(* Logix 5000 project; controller MV vendor 1 type 14 code 217 rev 31.11; software revision 31.00; part 8 of 53 *)
(* tags used below, declared in another part *)
   CWD : CHECKWORD_FLAGS;
   MC_B240 : INT[255];   // CH1 RN PMP Channel 1 return pum p drive flags
   MC_B242 : INT[255];   // CH1 ROUTE Channel 1 route requ est flags
   MC_bit_returned : BOOL;
   MC_CH1_DR1 : PlantItem;   // CH1_DR1
   MC_CH1_DR2 : PlantItem;   // CH1_DR2
   MC_CH1_DT1 : PlantItem;   // CH1_DT1
   MC_CH1_DT2 : PlantItem;   // CH1_DT2
   MC_CH1_R1 : PlantItem;   // CH1_R1
   MC_CH1_R1R : PlantItem;   // CH1_R1R
   MC_CH1_R2 : PlantItem;   // CH1_R2
   MC_CH1_R2R : PlantItem;   // CH1_R2R
   MC_CH1_R3 : PlantItem;   // CH1_R3
   MC_CH1_R3R : PlantItem;   // CH1_R3R
   MC_CH1_R4 : PlantItem;   // CH1_R4
   MC_CH1_R4R : PlantItem;   // CH1_R4R
   MC_CH1_R5 : PlantItem;   // CH1_R5
   MC_CH1_R5R : PlantItem;   // CH1_R5R
   MC_CH1_R6 : PlantItem;   // CH1_R6
   MC_CH1_R6R : PlantItem;   // CH1_R6R
   MC_CH1_T105_2_ACC : DINT;
   MC_data_file_value_to_move : DINT;
   MC_N10 : INT[255];   // SETTINGS
   MC_N100 : INT[255];   // C1_PLC Channel 1 PLC data
   MC_N100_29_0_Storagebit : BOOL;
   MC_N102 : INT[255];   // CH1 PROG Channel 1 CIP progra m
   MC_N104 : INT[255];   // CH1 REPORT Channel 1 CIP report file
   MC_N112 : INT[255];   // FVR DATA Data read from FV ro uting PLC
   MC_N113 : INT[255];   // MVR DATA Data read from MV ro uting PLC
   MC_N114 : INT[255];   // YP DATA
   MC_N200 : INT[255];   // CHK_WORK Plant item fault che cking work area
   MC_N7 : INT[255];   // INTEGER
   MC_P1 : PlantItem;   // P1
   MC_PX_100 : PlantItem;   // PX_100
   MC_PX_101 : PlantItem;   // PX_101
   MC_T105 : TIMER[255];   // CH1 TIMERS Channel 1 timers
   MC_T4 : TIMER[255];   // TIMER
(* MC_Common, continued *)

ROUTINE MC_CH1_GLOBL_105   (* ladder *)
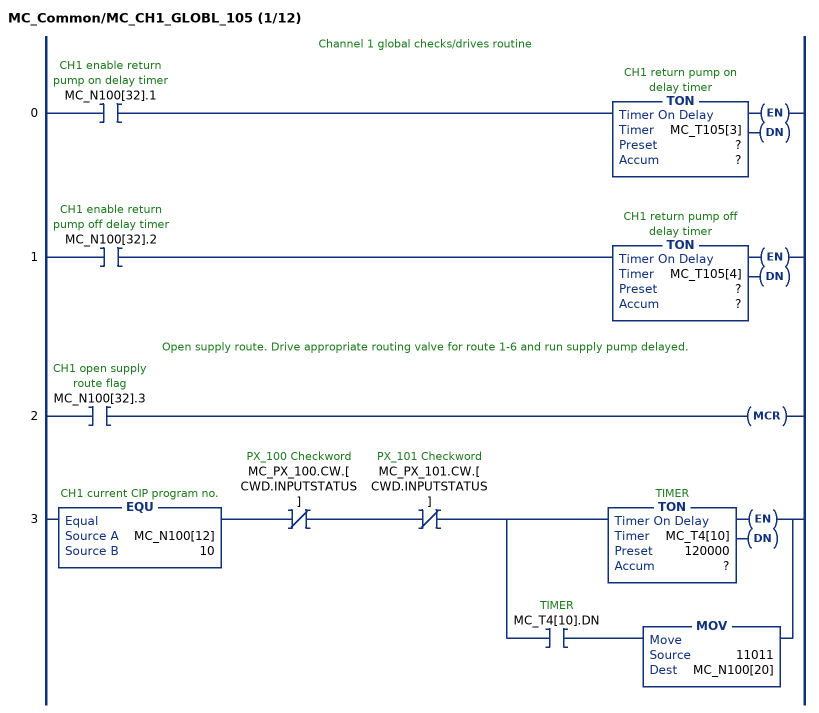
   // Channel 1 global checks/drives routine
   0: XIC(MC_N100[32].1)TON(MC_T105[3],?,?);
   1: XIC(MC_N100[32].2)TON(MC_T105[4],?,?);
   // Open supply route. Drive appropriate routing valve for route 1-6 and run supply pump delayed.
   2: XIC(MC_N100[32].3)MCR();
   3: EQU(MC_N100[12],10)XIO(MC_PX_100.CW.[CWD.INPUTSTATUS])XIO(MC_PX_101.CW.[CWD.INPUTSTATUS])[TON(MC_T4[10],?,?) ,XIC(MC_T4[10].DN) MOV(11011,MC_N100[20]) ];
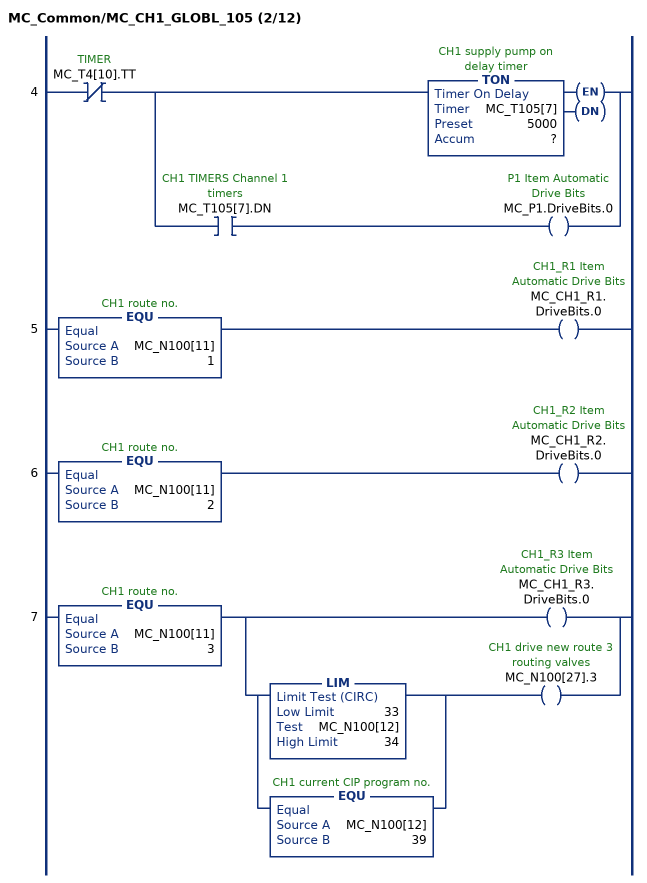
   4: XIO(MC_T4[10].TT)[TON(MC_T105[7],?,?) ,XIC(MC_T105[7].DN) OTE(MC_P1.DriveBits.0) ];
   5: EQU(MC_N100[11],1)OTE(MC_CH1_R1.DriveBits.0);
   6: EQU(MC_N100[11],2)OTE(MC_CH1_R2.DriveBits.0);
   7: EQU(MC_N100[11],3)[OTE(MC_CH1_R3.DriveBits.0) ,[LIM(33,MC_N100[12],34) ,EQU(MC_N100[12],39) ] OTE(MC_N100[27].3) ];
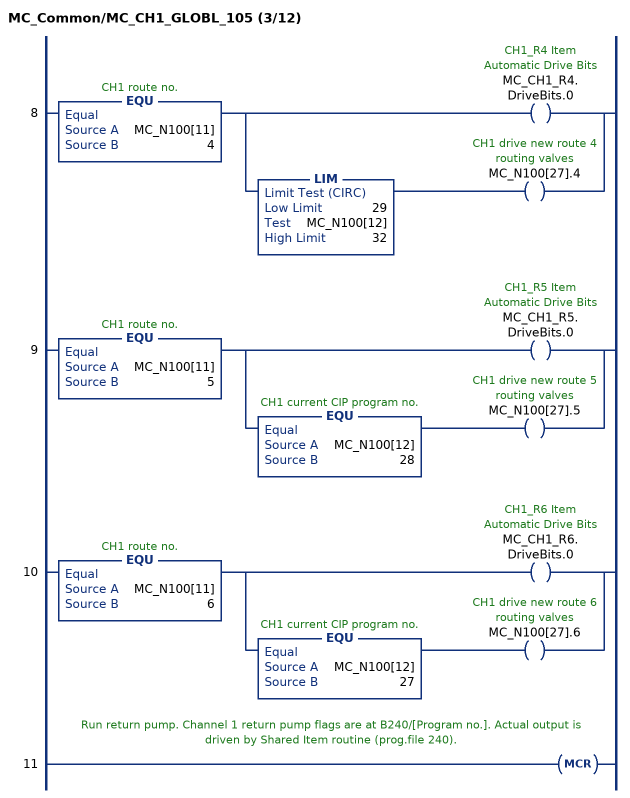
   8: EQU(MC_N100[11],4)[OTE(MC_CH1_R4.DriveBits.0) ,LIM(29,MC_N100[12],32) OTE(MC_N100[27].4) ];
   9: EQU(MC_N100[11],5)[OTE(MC_CH1_R5.DriveBits.0) ,EQU(MC_N100[12],28) OTE(MC_N100[27].5) ];
   10: EQU(MC_N100[11],6)[OTE(MC_CH1_R6.DriveBits.0) ,EQU(MC_N100[12],27) OTE(MC_N100[27].6) ];
   // Run return pump. Channel 1 return pump flags are at B240/[Program no.]. Actual output is driven by Shared Item routine (prog.file 240).
   11: MCR();
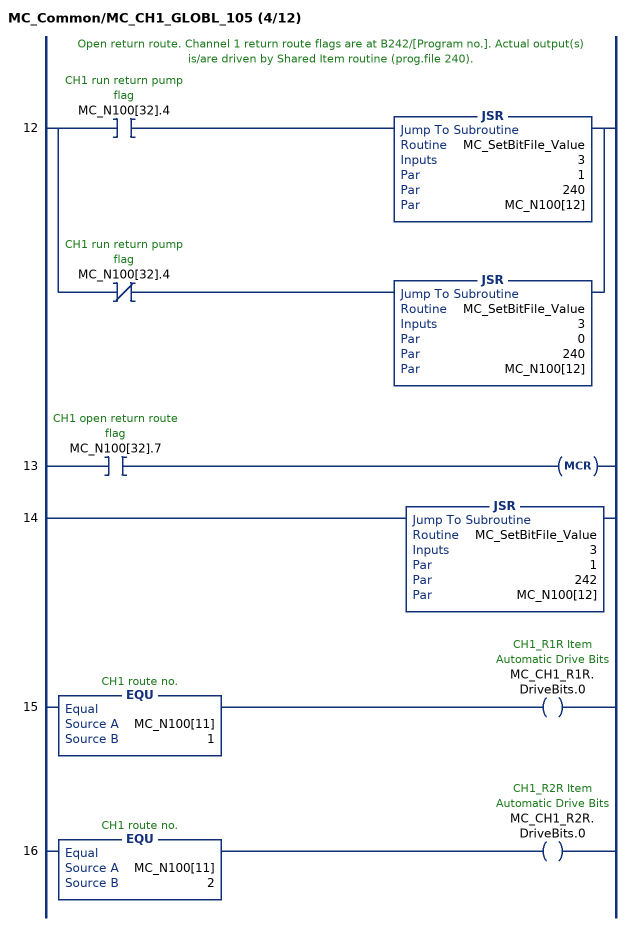
   // Open return route. Channel 1 return route flags are at B242/[Program no.]. Actual output(s) is/are driven by Shared Item routine (prog.file 240).
   12: [XIC(MC_N100[32].4) JSR(MC_SetBitFile_Value,3,1,240,MC_N100[12]) ,XIO(MC_N100[32].4) JSR(MC_SetBitFile_Value,3,0,240,MC_N100[12]) ];
   13: XIC(MC_N100[32].7)MCR();
   14: JSR(MC_SetBitFile_Value,3,1,242,MC_N100[12]);
   15: EQU(MC_N100[11],1)OTE(MC_CH1_R1R.DriveBits.0);
   16: EQU(MC_N100[11],2)OTE(MC_CH1_R2R.DriveBits.0);
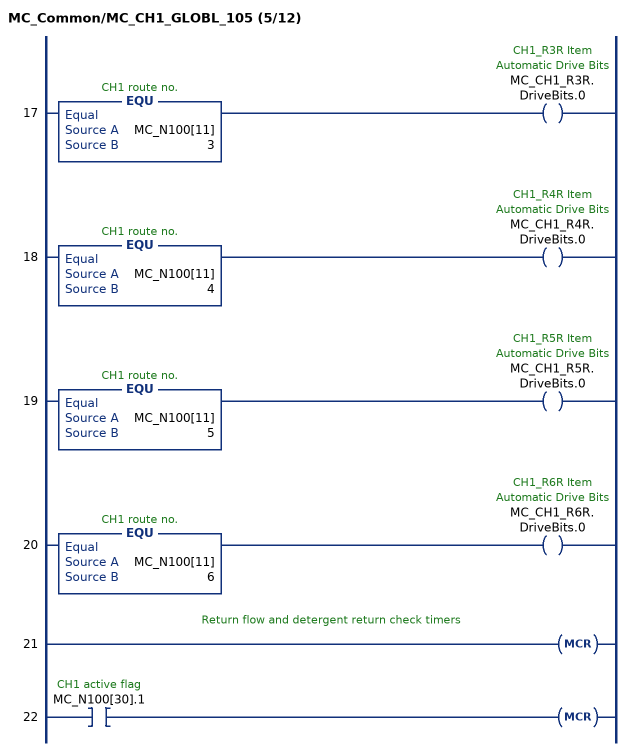
   17: EQU(MC_N100[11],3)OTE(MC_CH1_R3R.DriveBits.0);
   18: EQU(MC_N100[11],4)OTE(MC_CH1_R4R.DriveBits.0);
   19: EQU(MC_N100[11],5)OTE(MC_CH1_R5R.DriveBits.0);
   20: EQU(MC_N100[11],6)OTE(MC_CH1_R6R.DriveBits.0);
   // Return flow and detergent return check timers
   21: MCR();
   22: XIC(MC_N100[30].1)MCR();
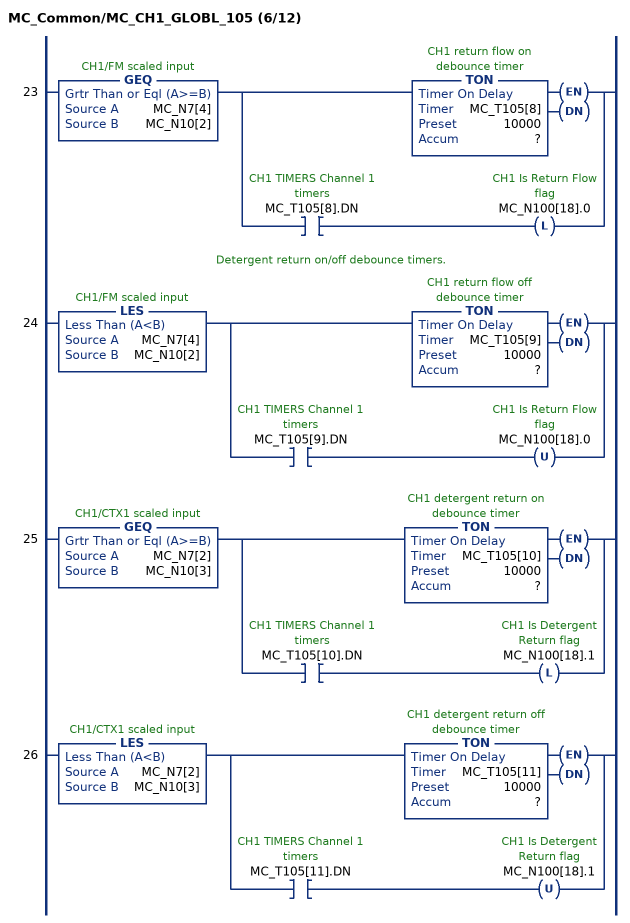
   23: GEQ(MC_N7[4],MC_N10[2])[TON(MC_T105[8],?,?) ,XIC(MC_T105[8].DN) OTL(MC_N100[18].0) ];
   // Detergent return on/off debounce timers.
   24: LES(MC_N7[4],MC_N10[2])[TON(MC_T105[9],?,?) ,XIC(MC_T105[9].DN) OTU(MC_N100[18].0) ];
   25: GEQ(MC_N7[2],MC_N10[3])[TON(MC_T105[10],?,?) ,XIC(MC_T105[10].DN) OTL(MC_N100[18].1) ];
   26: LES(MC_N7[2],MC_N10[3])[TON(MC_T105[11],?,?) ,XIC(MC_T105[11].DN) OTU(MC_N100[18].1) ];
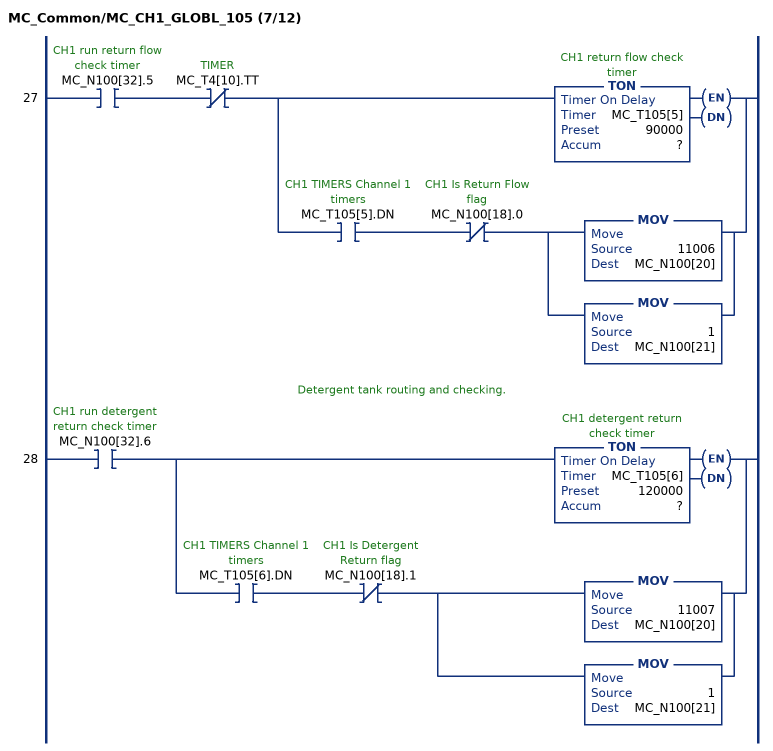
   27: XIC(MC_N100[32].5)XIO(MC_T4[10].TT)[TON(MC_T105[5],?,?) ,XIC(MC_T105[5].DN) XIO(MC_N100[18].0) [MOV(11006,MC_N100[20]) ,MOV(1,MC_N100[21]) ] ];
   // Detergent tank routing and checking.
   28: XIC(MC_N100[32].6)[TON(MC_T105[6],?,?) ,XIC(MC_T105[6].DN) XIO(MC_N100[18].1) [MOV(11007,MC_N100[20]) ,MOV(1,MC_N100[21]) ] ];
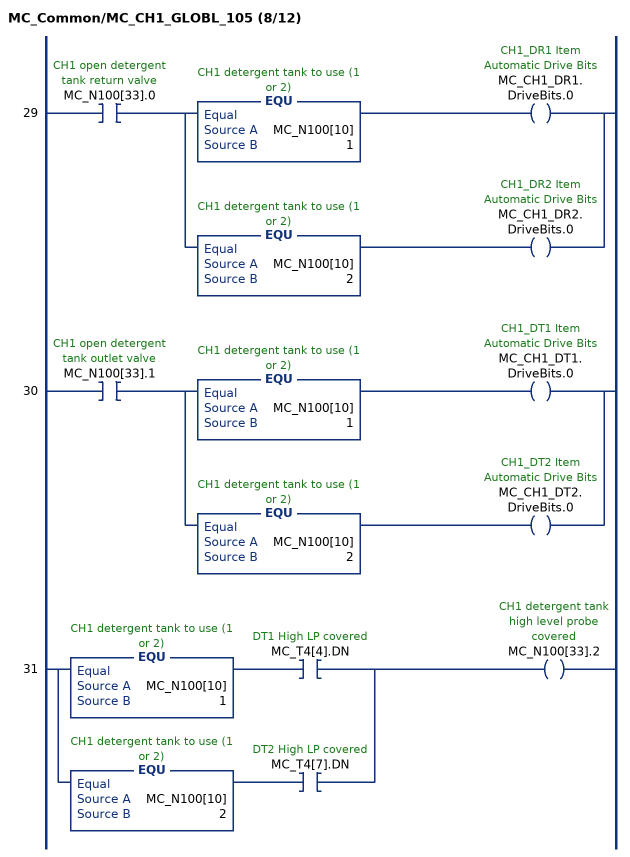
   29: XIC(MC_N100[33].0)[EQU(MC_N100[10],1) OTE(MC_CH1_DR1.DriveBits.0) ,EQU(MC_N100[10],2) OTE(MC_CH1_DR2.DriveBits.0) ];
   30: XIC(MC_N100[33].1)[EQU(MC_N100[10],1) OTE(MC_CH1_DT1.DriveBits.0) ,EQU(MC_N100[10],2) OTE(MC_CH1_DT2.DriveBits.0) ];
   31: [EQU(MC_N100[10],1) XIC(MC_T4[4].DN) ,EQU(MC_N100[10],2) XIC(MC_T4[7].DN) ]OTE(MC_N100[33].2);
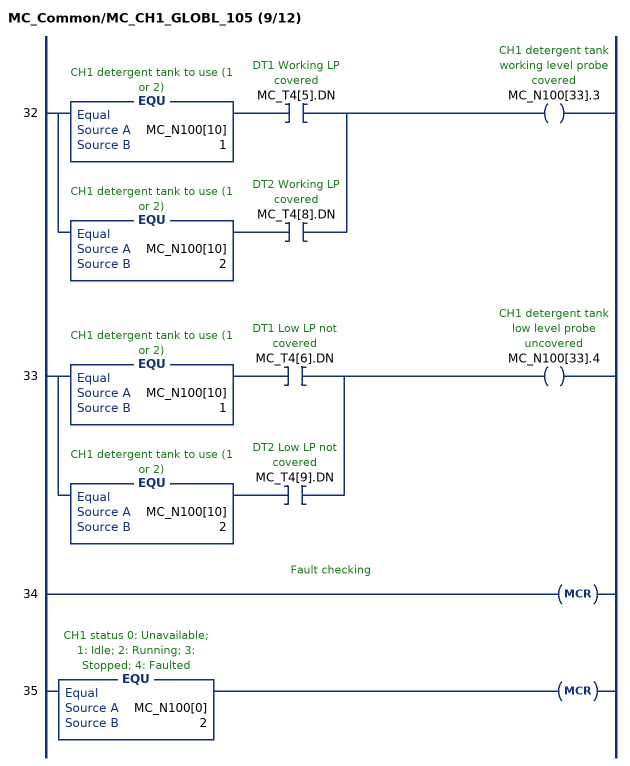
   32: [EQU(MC_N100[10],1) XIC(MC_T4[5].DN) ,EQU(MC_N100[10],2) XIC(MC_T4[8].DN) ]OTE(MC_N100[33].3);
   33: [EQU(MC_N100[10],1) XIC(MC_T4[6].DN) ,EQU(MC_N100[10],2) XIC(MC_T4[9].DN) ]OTE(MC_N100[33].4);
   // Fault checking
   34: MCR();
   35: EQU(MC_N100[0],2)MCR();
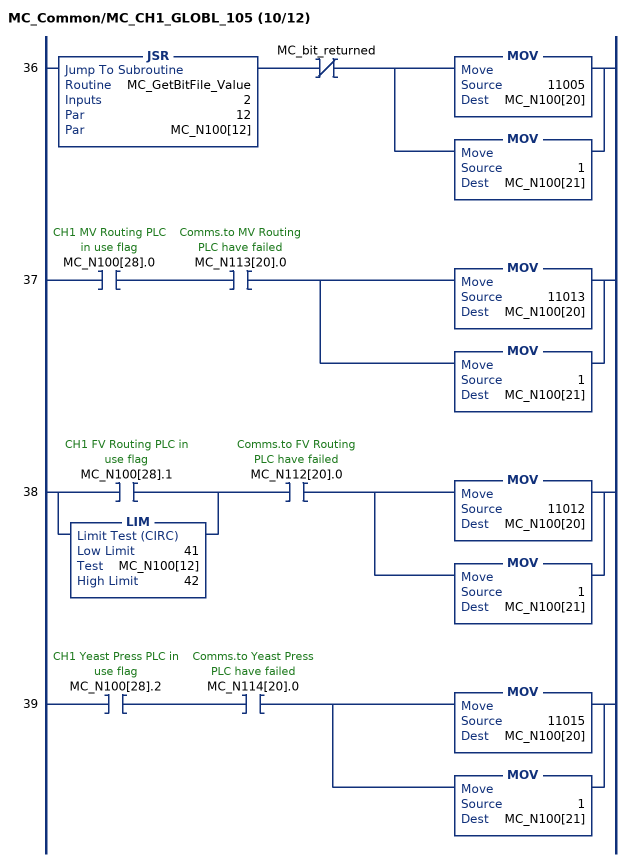
   36: JSR(MC_GetBitFile_Value,2,12,MC_N100[12])XIO(MC_bit_returned)[MOV(11005,MC_N100[20]) ,MOV(1,MC_N100[21]) ];
   37: XIC(MC_N100[28].0)XIC(MC_N113[20].0)[MOV(11013,MC_N100[20]) ,MOV(1,MC_N100[21]) ];
   38: [XIC(MC_N100[28].1) ,LIM(41,MC_N100[12],42) ]XIC(MC_N112[20].0)[MOV(11012,MC_N100[20]) ,MOV(1,MC_N100[21]) ];
   39: XIC(MC_N100[28].2)XIC(MC_N114[20].0)[MOV(11015,MC_N100[20]) ,MOV(1,MC_N100[21]) ];
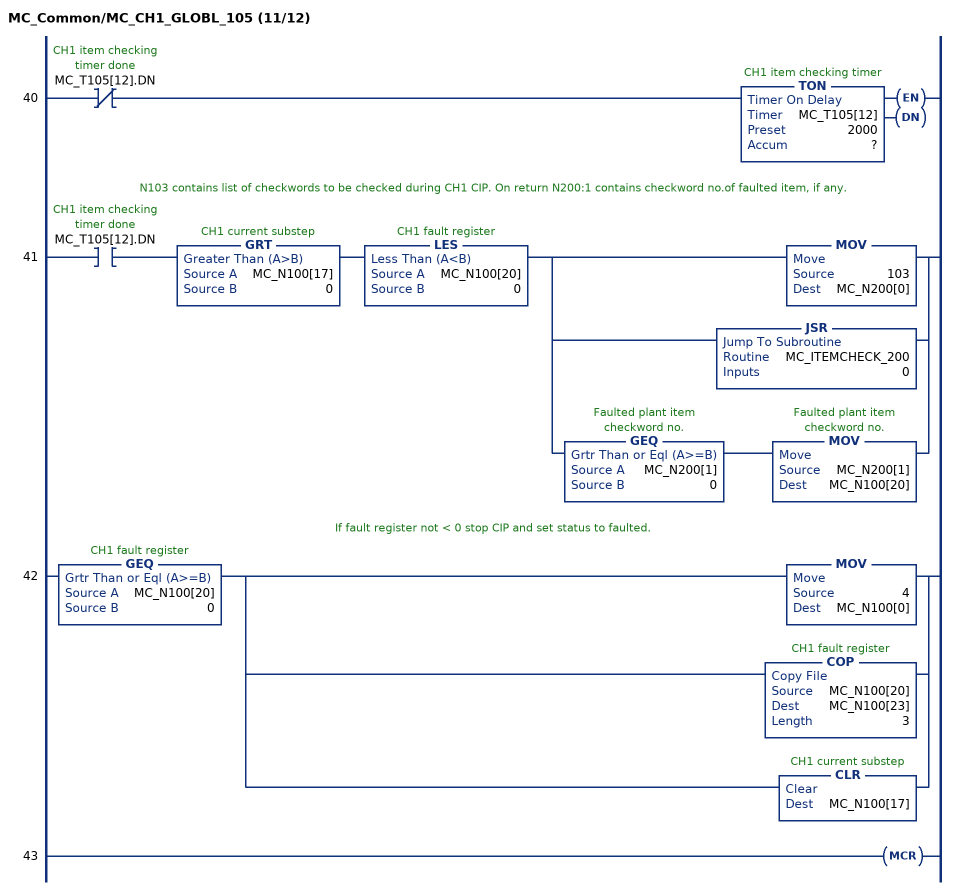
   40: XIO(MC_T105[12].DN)TON(MC_T105[12],?,?);
   // N103 contains list of checkwords to be checked during CH1 CIP. On return N200:1 contains checkword no.of faulted item, if any.
   41: XIC(MC_T105[12].DN)GRT(MC_N100[17],0)LES(MC_N100[20],0)[MOV(103,MC_N200[0]) ,JSR(MC_ITEMCHECK_200,0) ,GEQ(MC_N200[1],0) MOV(MC_N200[1],MC_N100[20]) ];
   // If fault register not < 0 stop CIP and set status to faulted.
   42: GEQ(MC_N100[20],0)[MOV(4,MC_N100[0]) ,COP(MC_N100[20],MC_N100[23],3) ,CLR(MC_N100[17]) ];
   43: MCR();
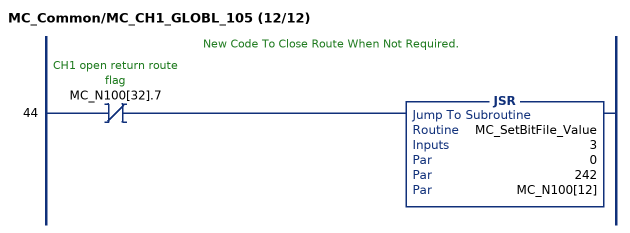
   // New Code To Close Route When Not Required.
   44: XIO(MC_N100[32].7)JSR(MC_SetBitFile_Value,3,0,242,MC_N100[12]);
END_ROUTINE

ROUTINE MC_CH1_MCP_100   (* ladder *)
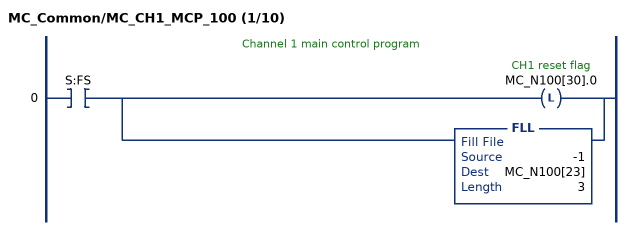
   // Channel 1 main control program
   0: XIC(S:FS)[OTL(MC_N100[30].0) ,FLL(-1,MC_N100[23],3) ];
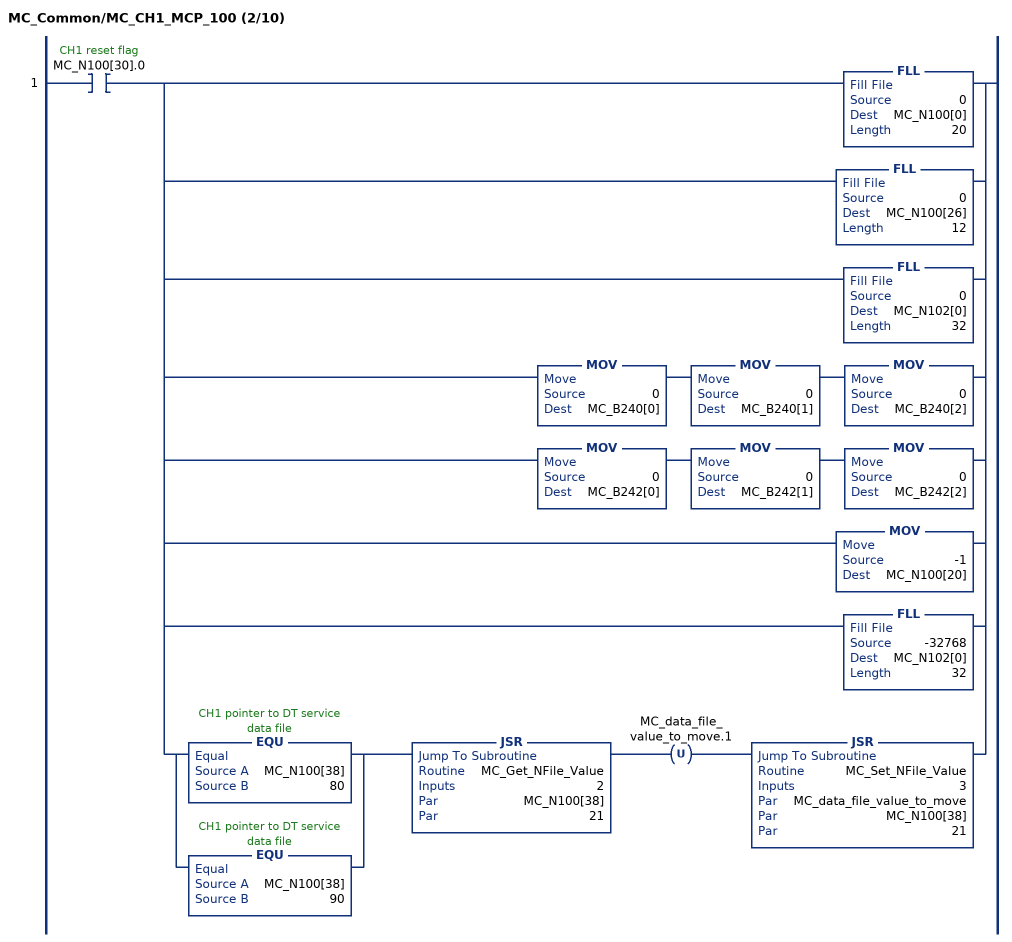
   1: XIC(MC_N100[30].0)[FLL(0,MC_N100[0],20) ,FLL(0,MC_N100[26],12) ,FLL(0,MC_N102[0],32) ,MOV(0,MC_B240[0]) MOV(0,MC_B240[1]) MOV(0,MC_B240[2]) ,MOV(0,MC_B242[0]) MOV(0,MC_B242[1]) MOV(0,MC_B242[2]) ,MOV(-1,MC_N100[20]) ,FLL(-32768,MC_N102[0],32) ,[EQU(MC_N100[38],80) ,EQU(MC_N100[38],90) ] JSR(MC_Get_NFile_Value,2,MC_N100[38],21) OTU(MC_data_file_value_to_move.1) JSR(MC_Set_NFile_Value,3,MC_data_file_value_to_move,MC_N100[38],21) ];
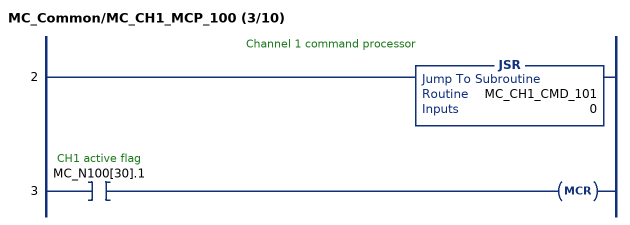
   // Channel 1 command processor
   2: JSR(MC_CH1_CMD_101,0);
   3: XIC(MC_N100[30].1)MCR();
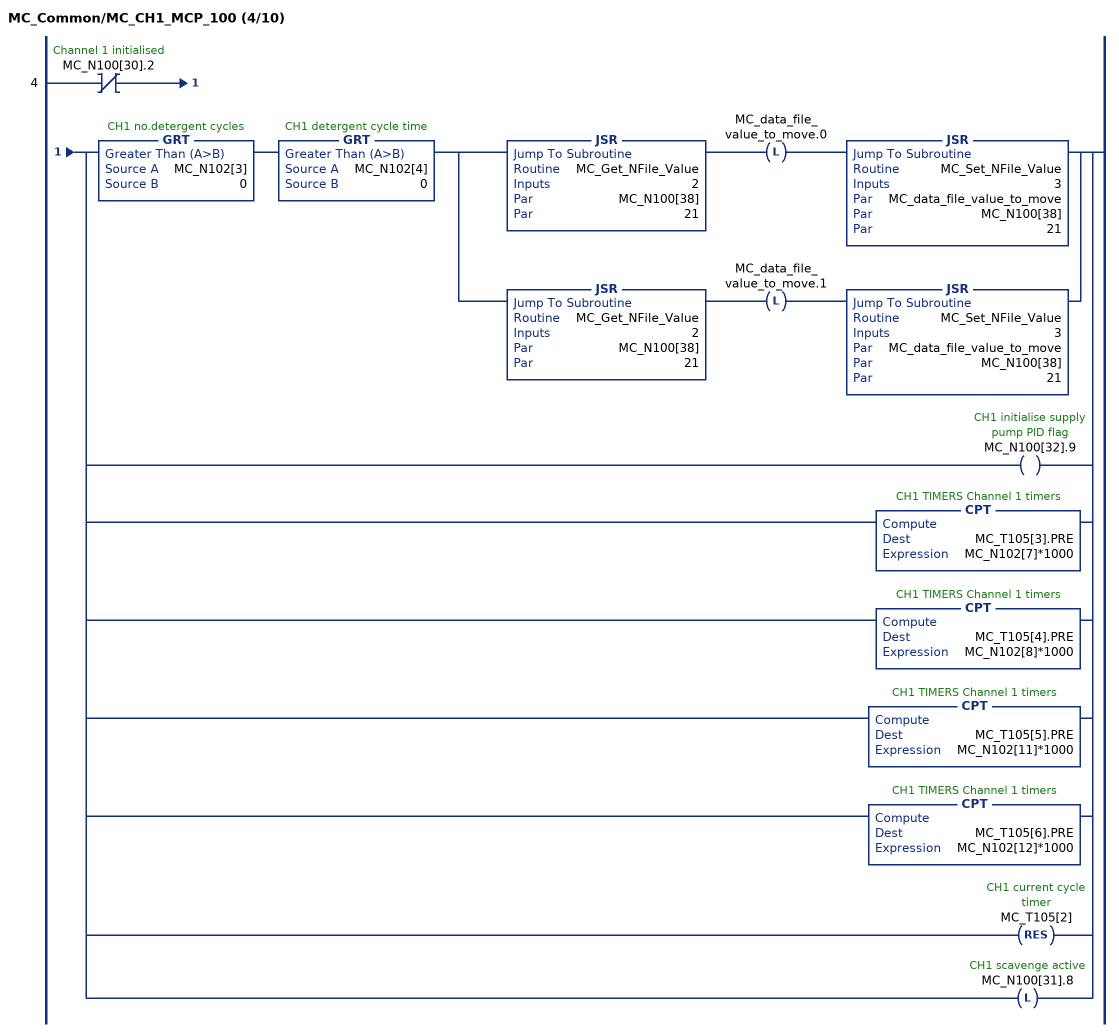
   4: XIO(MC_N100[30].2)[GRT(MC_N102[3],0) GRT(MC_N102[4],0) [JSR(MC_Get_NFile_Value,2,MC_N100[38],21) OTL(MC_data_file_value_to_move.0) JSR(MC_Set_NFile_Value,3,MC_data_file_value_to_move,MC_N100[38],21) ,JSR(MC_Get_NFile_Value,2,MC_N100[38],21) OTL(MC_data_file_value_to_move.1) JSR(MC_Set_NFile_Value,3,MC_data_file_value_to_move,MC_N100[38],21) ] ,OTE(MC_N100[32].9) ,[CPT(MC_T105[3].PRE,MC_N102[7]*1000) ,CPT(MC_T105[4].PRE,MC_N102[8]*1000) ,CPT(MC_T105[5].PRE,MC_N102[11]*1000) ,CPT(MC_T105[6].PRE,MC_N102[12]*1000) ,RES(MC_T105[2]) ,OTL(MC_N100[31].8) ] ];
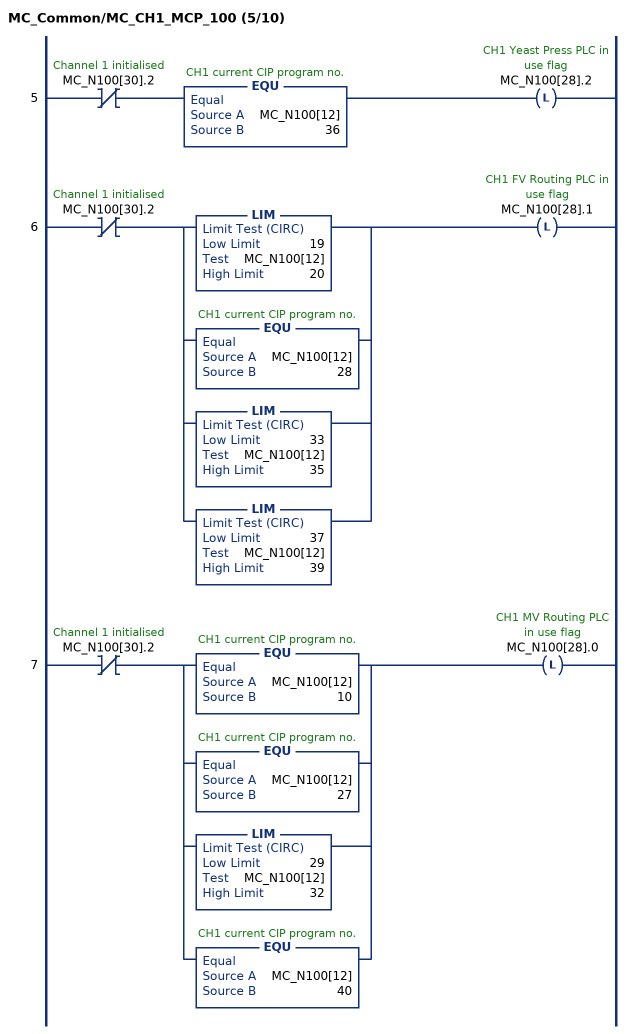
   5: XIO(MC_N100[30].2)EQU(MC_N100[12],36)OTL(MC_N100[28].2);
   6: XIO(MC_N100[30].2)[LIM(19,MC_N100[12],20) ,EQU(MC_N100[12],28) ,LIM(33,MC_N100[12],35) ,LIM(37,MC_N100[12],39) ]OTL(MC_N100[28].1);
   7: XIO(MC_N100[30].2)[EQU(MC_N100[12],10) ,EQU(MC_N100[12],27) ,LIM(29,MC_N100[12],32) ,EQU(MC_N100[12],40) ]OTL(MC_N100[28].0);
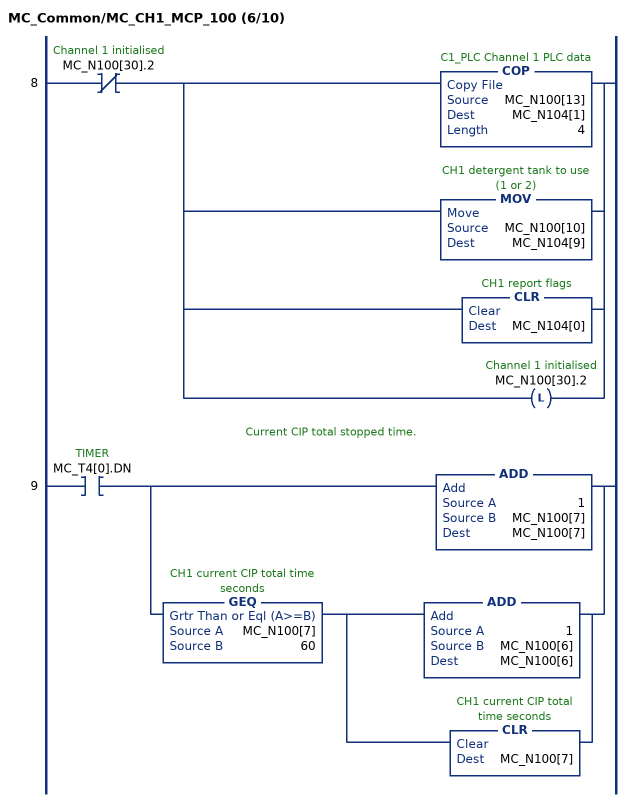
   8: XIO(MC_N100[30].2)[COP(MC_N100[13],MC_N104[1],4) ,MOV(MC_N100[10],MC_N104[9]) ,CLR(MC_N104[0]) ,OTL(MC_N100[30].2) ];
   // Current CIP total stopped time.
   9: XIC(MC_T4[0].DN)[ADD(1,MC_N100[7],MC_N100[7]) ,GEQ(MC_N100[7],60) [ADD(1,MC_N100[6],MC_N100[6]) ,CLR(MC_N100[7]) ] ];
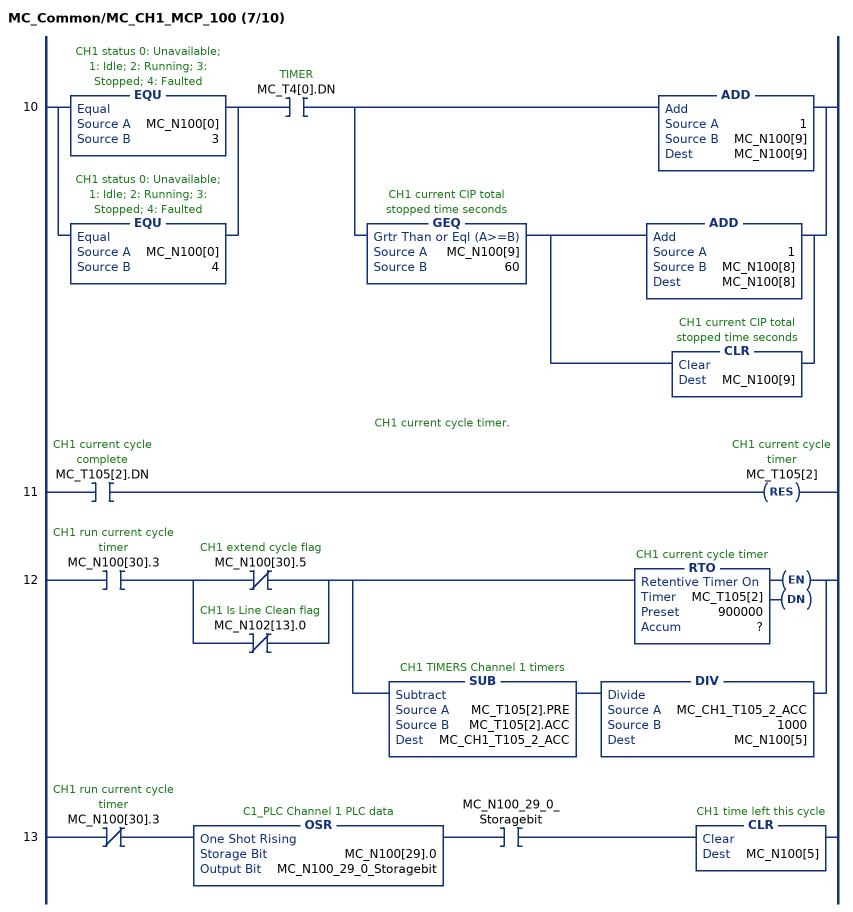
   10: [EQU(MC_N100[0],3) ,EQU(MC_N100[0],4) ]XIC(MC_T4[0].DN)[ADD(1,MC_N100[9],MC_N100[9]) ,GEQ(MC_N100[9],60) [ADD(1,MC_N100[8],MC_N100[8]) ,CLR(MC_N100[9]) ] ];
   // CH1 current cycle timer.
   11: XIC(MC_T105[2].DN)RES(MC_T105[2]);
   12: XIC(MC_N100[30].3)[XIO(MC_N100[30].5) ,XIO(MC_N102[13].0) ][RTO(MC_T105[2],?,?) ,SUB(MC_T105[2].PRE,MC_T105[2].ACC,MC_CH1_T105_2_ACC) DIV(MC_CH1_T105_2_ACC,1000,MC_N100[5]) ];
   13: XIO(MC_N100[30].3)OSR(MC_N100[29].0,MC_N100_29_0_Storagebit)XIC(MC_N100_29_0_Storagebit)CLR(MC_N100[5]);
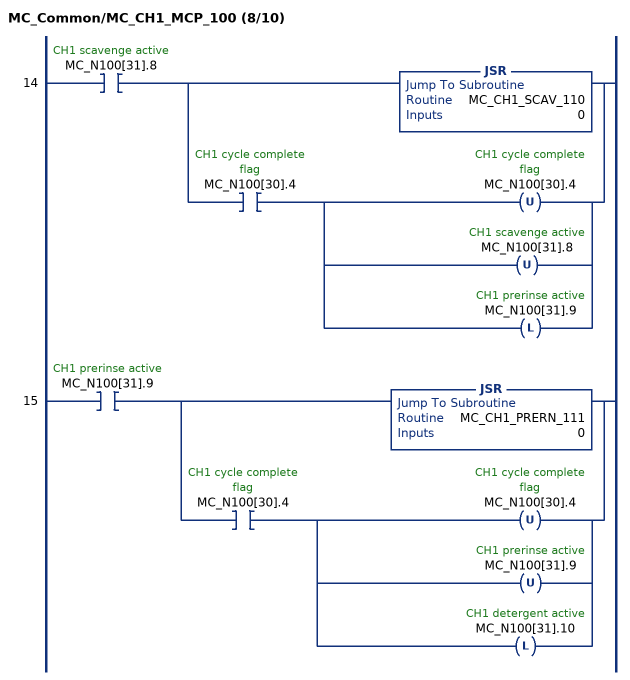
   14: XIC(MC_N100[31].8)[JSR(MC_CH1_SCAV_110,0) ,XIC(MC_N100[30].4) [OTU(MC_N100[30].4) ,OTU(MC_N100[31].8) ,OTL(MC_N100[31].9) ] ];
   15: XIC(MC_N100[31].9)[JSR(MC_CH1_PRERN_111,0) ,XIC(MC_N100[30].4) [OTU(MC_N100[30].4) ,OTU(MC_N100[31].9) ,OTL(MC_N100[31].10) ] ];
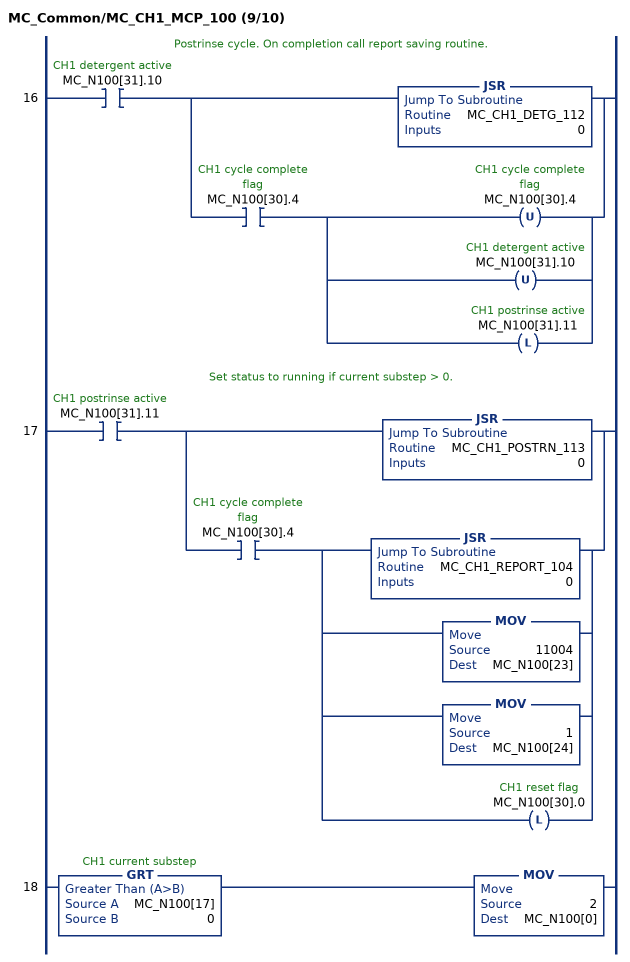
   // Postrinse cycle. On completion call report saving routine.
   16: XIC(MC_N100[31].10)[JSR(MC_CH1_DETG_112,0) ,XIC(MC_N100[30].4) [OTU(MC_N100[30].4) ,OTU(MC_N100[31].10) ,OTL(MC_N100[31].11) ] ];
   // Set status to running if current substep > 0.
   17: XIC(MC_N100[31].11)[JSR(MC_CH1_POSTRN_113,0) ,XIC(MC_N100[30].4) [JSR(MC_CH1_REPORT_104,0) ,MOV(11004,MC_N100[23]) ,MOV(1,MC_N100[24]) ,OTL(MC_N100[30].0) ] ];
   18: GRT(MC_N100[17],0)MOV(2,MC_N100[0]);
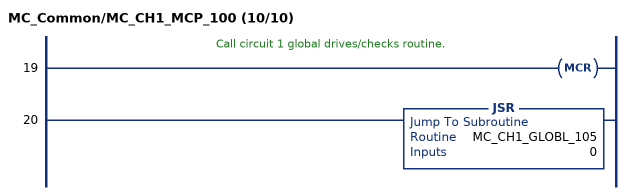
   // Call circuit 1 global drives/checks routine.
   19: MCR();
   20: JSR(MC_CH1_GLOBL_105,0);
END_ROUTINE
